DATA_BLOCK "LANGUAGE"   // DB4
TITLE = LANGUAGE
{ S7_Optimized_Access := 'FALSE' }
AUTHOR : oscat
FAMILY : CONSTANT
NAME : DBLANG
VERSION : 1.2
   VAR
      DEFAULT : Int := 1;   // 1=english, 2=german, 3=french
      LMAX : Int := 3;
      WEEKDAYS : Array[1..3, 1..7] of String[10];
      WEEKDAYS2 : Array[1..3, 1..7] of String[2];
      MONTHS : Array[1..3, 1..12] of String[10];
      MONTHS3 : Array[1..3, 1..12] of String[3];
      DIRS : Array[1..3, 0..15] of String[3];
   END_VAR
BEGIN
   WEEKDAYS[1,1] := 'Monday';
   WEEKDAYS[1,2] := 'Tuesday';
   WEEKDAYS[1,3] := 'Wednesday';
   WEEKDAYS[1,4] := 'Thursday';
   WEEKDAYS[1,5] := 'Friday';
   WEEKDAYS[1,6] := 'Saturday';
   WEEKDAYS[1,7] := 'Sunday';
   WEEKDAYS[2,1] := 'Montag';
   WEEKDAYS[2,2] := 'Dienstag';
   WEEKDAYS[2,3] := 'Mittwoch';
   WEEKDAYS[2,4] := 'Donnerstag';
   WEEKDAYS[2,5] := 'Freitag';
   WEEKDAYS[2,6] := 'Samstag';
   WEEKDAYS[2,7] := 'Sonntag';
   WEEKDAYS[3,1] := 'Lundi';
   WEEKDAYS[3,2] := 'Mardi';
   WEEKDAYS[3,3] := 'Mercredi';
   WEEKDAYS[3,4] := 'Jeudi';
   WEEKDAYS[3,5] := 'Vendredi';
   WEEKDAYS[3,6] := 'Samedi';
   WEEKDAYS[3,7] := 'Dimanche';
   WEEKDAYS2[1,1] := 'Mo';
   WEEKDAYS2[1,2] := 'Tu';
   WEEKDAYS2[1,3] := 'We';
   WEEKDAYS2[1,4] := 'Th';
   WEEKDAYS2[1,5] := 'Fr';
   WEEKDAYS2[1,6] := 'Sa';
   WEEKDAYS2[1,7] := 'Su';
   WEEKDAYS2[2,1] := 'Mo';
   WEEKDAYS2[2,2] := 'Di';
   WEEKDAYS2[2,3] := 'Mi';
   WEEKDAYS2[2,4] := 'Do';
   WEEKDAYS2[2,5] := 'Fr';
   WEEKDAYS2[2,6] := 'Sa';
   WEEKDAYS2[2,7] := 'So';
   WEEKDAYS2[3,1] := 'Lu';
   WEEKDAYS2[3,2] := 'Ma';
   WEEKDAYS2[3,3] := 'Me';
   WEEKDAYS2[3,4] := 'Je';
   WEEKDAYS2[3,5] := 'Ve';
   WEEKDAYS2[3,6] := 'Sa';
   WEEKDAYS2[3,7] := 'Di';
   MONTHS[1,1] := 'January';
   MONTHS[1,2] := 'February';
   MONTHS[1,3] := 'March';
   MONTHS[1,4] := 'April';
   MONTHS[1,5] := 'May';
   MONTHS[1,6] := 'June';
   MONTHS[1,7] := 'July';
   MONTHS[1,8] := 'August';
   MONTHS[1,9] := 'September';
   MONTHS[1,10] := 'October';
   MONTHS[1,11] := 'November';
   MONTHS[1,12] := 'December';
   MONTHS[2,1] := 'Januar';
   MONTHS[2,2] := 'Februar';
   MONTHS[2,3] := 'März';
   MONTHS[2,4] := 'April';
   MONTHS[2,5] := 'Mai';
   MONTHS[2,6] := 'Juni';
   MONTHS[2,7] := 'Juli';
   MONTHS[2,8] := 'August';
   MONTHS[2,9] := 'September';
   MONTHS[2,10] := 'Oktober';
   MONTHS[2,11] := 'November';
   MONTHS[2,12] := 'Dezember';
   MONTHS[3,1] := 'Janvier';
   MONTHS[3,2] := 'Février';
   MONTHS[3,3] := 'mars';
   MONTHS[3,4] := 'Avril';
   MONTHS[3,5] := 'Mai';
   MONTHS[3,6] := 'Juin';
   MONTHS[3,7] := 'Juillet';
   MONTHS[3,8] := 'Août';
   MONTHS[3,9] := 'Septembre';
   MONTHS[3,10] := 'Octobre';
   MONTHS[3,11] := 'Novembre';
   MONTHS[3,12] := 'Decembre';
   MONTHS3[1,1] := 'Jan';
   MONTHS3[1,2] := 'Feb';
   MONTHS3[1,3] := 'Mar';
   MONTHS3[1,4] := 'Apr';
   MONTHS3[1,5] := 'May';
   MONTHS3[1,6] := 'Jun';
   MONTHS3[1,7] := 'Jul';
   MONTHS3[1,8] := 'Aug';
   MONTHS3[1,9] := 'Sep';
   MONTHS3[1,10] := 'Oct';
   MONTHS3[1,11] := 'Nov';
   MONTHS3[1,12] := 'Dec';
   MONTHS3[2,1] := 'Jan';
   MONTHS3[2,2] := 'Feb';
   MONTHS3[2,3] := 'Mrz';
   MONTHS3[2,4] := 'Apr';
   MONTHS3[2,5] := 'Mai';
   MONTHS3[2,6] := 'Jun';
   MONTHS3[2,7] := 'Jul';
   MONTHS3[2,8] := 'Aug';
   MONTHS3[2,9] := 'Sep';
   MONTHS3[2,10] := 'Okt';
   MONTHS3[2,11] := 'Nov';
   MONTHS3[2,12] := 'Dez';
   MONTHS3[3,1] := 'Jan';
   MONTHS3[3,2] := 'Fev';
   MONTHS3[3,3] := 'Mar';
   MONTHS3[3,4] := 'Avr';
   MONTHS3[3,5] := 'Mai';
   MONTHS3[3,6] := 'Jun';
   MONTHS3[3,7] := 'Jul';
   MONTHS3[3,8] := 'Aou';
   MONTHS3[3,9] := 'Sep';
   MONTHS3[3,10] := 'Oct';
   MONTHS3[3,11] := 'Nov';
   MONTHS3[3,12] := 'Dec';
   DIRS[1,0] := 'N';
   DIRS[1,1] := 'NNE';
   DIRS[1,2] := 'NE';
   DIRS[1,3] := 'ENE';
   DIRS[1,4] := 'E';
   DIRS[1,5] := 'ESE';
   DIRS[1,6] := 'SE';
   DIRS[1,7] := 'SSE';
   DIRS[1,8] := 'S';
   DIRS[1,9] := 'SSW';
   DIRS[1,10] := 'SW';
   DIRS[1,11] := 'WSW';
   DIRS[1,12] := 'W';
   DIRS[1,13] := 'WNW';
   DIRS[1,14] := 'NW';
   DIRS[1,15] := 'NNW';
   DIRS[2,0] := 'N';
   DIRS[2,1] := 'NNO';
   DIRS[2,2] := 'NO';
   DIRS[2,3] := 'ONO';
   DIRS[2,4] := 'O';
   DIRS[2,5] := 'OSO';
   DIRS[2,6] := 'SO';
   DIRS[2,7] := 'SSO';
   DIRS[2,8] := 'S';
   DIRS[2,9] := 'SSW';
   DIRS[2,10] := 'SW';
   DIRS[2,11] := 'WSW';
   DIRS[2,12] := 'W';
   DIRS[2,13] := 'WNW';
   DIRS[2,14] := 'NW';
   DIRS[2,15] := 'NNW';
   DIRS[3,0] := 'N';
   DIRS[3,1] := 'NNO';
   DIRS[3,2] := 'NO';
   DIRS[3,3] := 'ONO';
   DIRS[3,4] := 'O';
   DIRS[3,5] := 'OSO';
   DIRS[3,6] := 'SO';
   DIRS[3,7] := 'SSO';
   DIRS[3,8] := 'S';
   DIRS[3,9] := 'SSW';
   DIRS[3,10] := 'SW';
   DIRS[3,11] := 'WSW';
   DIRS[3,12] := 'W';
   DIRS[3,13] := 'WNW';
   DIRS[3,14] := 'NW';
   DIRS[3,15] := 'NNW';
END_DATA_BLOCK

DATA_BLOCK "CONSTANTS"   // DB6
TITLE = CONSTANTS
{ S7_Optimized_Access := 'FALSE' }
AUTHOR : oscat
FAMILY : CONSTANT
NAME : CONSTANT
VERSION : 1.0
   VAR
      STRING_LENGTH : Int := 250;
      LIST_LENGTH : Int := 250;
   END_VAR
BEGIN
END_DATA_BLOCK

DATA_BLOCK "TEMP"   // DB7
TITLE = temporary Strings
{ S7_Optimized_Access := 'FALSE' }
AUTHOR : dalbi
FAMILY : xS7
NAME : DBTEMP
VERSION : 1.1
   VAR
      STR1 : String[254];
      STR2 : String[254];
      STR3 : String[254];
      TEMP : String[254];
   END_VAR
BEGIN
END_DATA_BLOCK

FUNCTION_BLOCK "MESSAGE_4R"   // FB34, SCL
TITLE = MESSAGE_4R
{ S7_Optimized_Access := 'FALSE' }
AUTHOR : hugo
FAMILY : STRINGS
NAME : MESSG4R
VERSION : 1.1
// this function generates a rotation meassage with up to 4 strings.
// on each rising edge of EN the next message in line will be displayed.
// when EN stays high longer then one cycle, the next message will be displayed automatically after the time T1 is elapsed.
// the output MX is the generated message and CX is a counter 0..3 signaling the current message displayed.
// the displayed messages are 0 .. MM.
// 
// uses: INC1 [FC53]
   VAR_INPUT
      M0 : String[254];
      M1 : String[254];
      M2 : String[254];
      M3 : String[254];
      MM : Int := 3;
      ENQ : Bool := TRUE;
      CLK : Bool := TRUE;
      T1 : Time := T#3S;
   END_VAR
   VAR_OUTPUT
      MX : String[254];
      MN : Int;
      TR : Bool;
   END_VAR
   VAR
      _timer : TON;
      edge : Bool;
   END_VAR
BEGIN


   (* check for rising edge on EN *)
   #TR := FALSE;
   IF #ENQ THEN
       IF (NOT #edge AND #CLK) OR #_timer.Q THEN
               #MN := "INC1"(N:=#MM,X:=#MN);
               #TR := TRUE;
               #_timer.IN := FALSE;
               CASE #MN OF
                   0 : #MX BLKMOV #M0;
                   1 : #MX BLKMOV #M1;
                   2 : #MX BLKMOV #M2;
                   3 : #MX BLKMOV #M3;
               END_CASE;
       END_IF;
       #edge := #CLK;
       #_timer( IN := #CLK, PT := #T1);
   ELSE
       #MX := '';
       #MN := 0;
   END_IF;




   (* revision history
   hm  8. oct. 2008    rev 1.0
       original version

   hm  27. oct. 2008   rev 1.1
       changed _INC to INC1

   *)
END_FUNCTION_BLOCK

FUNCTION_BLOCK "MESSAGE_8"   // FB35, SCL
TITLE = MESSAGE_8
{ S7_Optimized_Access := 'FALSE' }
AUTHOR : hugo
FAMILY : STRINGS
NAME : MESSAGE8
VERSION : 1.1
// this function generates one out of 4 messages specified by S1 .. S8.
// the selected message will be presented at the output M.
// In1 has higher priority then In2 which has higher priority then IN3 and in8 has the lowest priority.
   VAR_INPUT
      IN1 : Bool;
      IN2 : Bool;
      IN3 : Bool;
      IN4 : Bool;
      IN5 : Bool;
      IN6 : Bool;
      IN7 : Bool;
      IN8 : Bool;
      S1 : String[254];
      S2 : String[254];
      S3 : String[254];
      S4 : String[254];
      S5 : String[254];
      S6 : String[254];
      S7 : String[254];
      S8 : String[254];
   END_VAR
   VAR_OUTPUT
      "M" : String[254];
   END_VAR
BEGIN


     (* check if an alarm is present if yes set the output M otherwise clear M *)
     IF #IN1 THEN
       #"M" BLKMOV #S1;
     ELSIF #IN2 THEN
       #"M" BLKMOV #S2;
     ELSIF #IN3 THEN
       #"M" BLKMOV #S3;
     ELSIF #IN4 THEN
       #"M" BLKMOV #S4;
     ELSIF #IN5 THEN
       #"M" BLKMOV #S5;
     ELSIF #IN6 THEN
       #"M" BLKMOV #S6;
     ELSIF #IN7 THEN
       #"M" BLKMOV #S7;
     ELSIF #IN8 THEN
       #"M" BLKMOV #S8;
     ELSE
       #"M" := '';
     END_IF;

   (* revision history
   hm  26.12.2007      rev 1.0
       original version

   hm  29. mar. 2008   rev 1.1
       changed STRING to STRING(STRING_LENGTH)
   *)
END_FUNCTION_BLOCK

FUNCTION_BLOCK "TICKER"   // FB36, SCL
TITLE = TICKER
{ S7_Optimized_Access := 'FALSE' }
AUTHOR : hugo
FAMILY : STRINGS
NAME : TICKER
VERSION : 1.2
// Ticker sends a substring of text with length N every TD Milliseconds to generate a ticker. 
//  
// uses: MID [FC26]
   VAR_INPUT
      N : Int;
      PT : Time;
   END_VAR
   VAR_OUTPUT
      Display : String[254];
   END_VAR
   VAR_IN_OUT
      Text : String[254];
   END_VAR
   VAR
      delay : TP;
      "step" : Int;
   END_VAR
   VAR_TEMP
      tText : String[254];
      _Text AT tText : Struct
         length : Byte;
         act_length : Byte;
         str : Array[1..254] of Byte;
      END_STRUCT;
   END_VAR
BEGIN


   #tText := #Text; 

   (* generate next ticker when delay is low *)
   IF #N < BYTE_TO_INT(#_Text.act_length) THEN
       IF NOT #delay.Q THEN
         (* increase step for next tick *)
         #"step" := #"step" + 1;
         IF #"step" > BYTE_TO_INT(#_Text.act_length) THEN #"step" := 1; END_IF;
         (* extract dispay from text *)
         #Display := MID(IN:=#tText,L:=#N,P:=#"step");
         (* set delay timer for next tick *)
         #delay(IN := TRUE, PT := #PT);
       ELSE;
         (* execute delay timer *)
         #delay.IN := FALSE;
       END_IF;
   ELSE
       #Display BLKMOV #tText;
   END_IF;


   (* revision history
   hm  4. dec. 2007    rev 1.0
       original version

   hm  15. dec. 2007   rev 1.1
       step now starts at 1 instaed of 0

   hm  29. mar. 2008   rev 1.2
       changed STRING to STRING(STRING_LENGTH)
   *)
END_FUNCTION_BLOCK

FUNCTION "INC1" : Int   // FC53, SCL
TITLE = INC1
{ S7_Optimized_Access := 'FALSE' }
AUTHOR : hugo
FAMILY : MATH
NAME : INC1
VERSION : 1.2
// This is a increment function which increments the variable X by 1 and if M is reached, it begins with 0 again.
// _inc1(3,X) will generate 0,1,2,3,0,1,.....
   VAR_INPUT
      X : Int;
      N : Int;
   END_VAR
BEGIN


   IF #X >= #N - 1 THEN
       #INC1 := 0;
   ELSE
       #INC1 := #X + 1;
   END_IF;


   (* this elegant version is 50% slower
   INC1 := X := (x + 1) MOD N;
   *)



   (* revision history
   hm  13. oct. 2008   rev 1.0
       original version

   hm  22. oct. 2008   rev 1.1
       added statement to return value for compatibility reasons

   hm  23. feb. 2009   rev 1.2
       when inc1 is called with X >= N inc will continue with 0
   *)
END_FUNCTION

FUNCTION "EXP10" : Real   // FC77, SCL
TITLE = EXP10
{ S7_Optimized_Access := 'FALSE' }
AUTHOR : hugo
FAMILY : MATH
NAME : exp10
VERSION : 1.0
// this function calculates the exponent to the basis 10
// exp10(3) = 1000
   VAR_INPUT
      X : Real;
   END_VAR
BEGIN


     #EXP10 := EXP(#X * 2.30258509299405);

   (* revision history
   hm  2. dec 2007    rev 1.0
     original version

   *)
END_FUNCTION

FUNCTION "EXPN" : Real   // FC78, SCL
TITLE = EXPN
{ S7_Optimized_Access := 'FALSE' }
AUTHOR : hugo
FAMILY : MATH
NAME : EXPN
VERSION : 1.2
// this function calculates X to the power of N (Y = X^N) whilke N is an integer
// especially on CPU's without a floating point unit this algorythm is about 30 times faster then the IEC standard EXPT() Function
   VAR_INPUT
      X : Real;
      N : Int;
   END_VAR
   VAR_TEMP
      tempN : Int;
      _tempN AT tempN : Array[0..15] of Bool;
      tempX : Real;
      sign : Bool;
   END_VAR
BEGIN


   #tempN := #N;
   #tempX := #X;

   #sign := #_tempN[7]; //N.15
   #tempN := ABS(#tempN);
   IF #_tempN[8] THEN #EXPN := #tempX; ELSE #EXPN := 1.0; END_IF;
   #tempN := WORD_TO_INT(SHR(IN:=INT_TO_WORD(#tempN),N:=1));
   WHILE #tempN > 0 DO
      #tempX := #tempX * #tempX;
      IF #_tempN[8] THEN #EXPN := #EXPN * #tempX; END_IF;
      #tempN := WORD_TO_INT(SHR(IN:=INT_TO_WORD(#tempN),N:=1));
   END_WHILE;
   IF #sign THEN #EXPN := 1.0 / #EXPN; END_IF;


   (* revision history
   hm  4. dec 2007 rev 1.0
       original version

   hm  22. oct. 2008   rev 1.1
       optimized code

   hm  10. mar. 2009   rev 1.2
       removed nested comments
       real constants updated to new systax using dot

   *)
END_FUNCTION

FUNCTION "DAY_OF_MONTH" : Int   // FC178, SCL
TITLE = DAY_OF_MONTH
{ S7_Optimized_Access := 'FALSE' }
AUTHOR : hugo
FAMILY : TIDT
NAME : DAYOMON
VERSION : 2.1
// returns the day OF month from any DATE
// 
// uses: DAY_OF_YEAR [FC180]
//       YEAR_BEGIN [FC217] 
//       YEAR_OF_DATE [FC219] 
//       LEAP_OF_DATE [FC193]
//       LEAP_YEAR [FC194]
   VAR_INPUT
      IDATE : Date;
   END_VAR
   VAR_TEMP
      leap : Int;
   END_VAR
BEGIN


   (* calculate the day in the year *)
   #DAY_OF_MONTH := "DAY_OF_YEAR"(#IDATE);
   (* leap will be set to one for a leap year *)
   #leap := BOOL_TO_INT("LEAP_OF_DATE"(#IDATE));
   (* if leap year deduct one from the days of the year *)
   #DAY_OF_MONTH := #DAY_OF_MONTH - #leap;
   (* search if we are in month december to march ? *)
   IF #DAY_OF_MONTH > "MTH_OFS9" THEN
       IF #DAY_OF_MONTH > "MTH_OFS11" THEN
           IF #DAY_OF_MONTH > "MTH_OFS12" THEN
               #DAY_OF_MONTH := #DAY_OF_MONTH - "MTH_OFS12";
           ELSE
               #DAY_OF_MONTH := #DAY_OF_MONTH - "MTH_OFS11";
           END_IF;
       ELSE
           IF #DAY_OF_MONTH > "MTH_OFS10" THEN
               #DAY_OF_MONTH := #DAY_OF_MONTH - "MTH_OFS10";
           ELSE
               #DAY_OF_MONTH := #DAY_OF_MONTH - "MTH_OFS9";
           END_IF;
       END_IF;
   ELSIF #DAY_OF_MONTH > "MTH_OFS5" THEN
       IF #DAY_OF_MONTH > "MTH_OFS7" THEN
           IF #DAY_OF_MONTH > "MTH_OFS8" THEN
               #DAY_OF_MONTH := #DAY_OF_MONTH - "MTH_OFS8";
           ELSE
               #DAY_OF_MONTH := #DAY_OF_MONTH - "MTH_OFS7";
           END_IF;
       ELSE
           IF #DAY_OF_MONTH > "MTH_OFS6" THEN
               #DAY_OF_MONTH := #DAY_OF_MONTH - "MTH_OFS6";
           ELSE
               #DAY_OF_MONTH := #DAY_OF_MONTH - "MTH_OFS5";
           END_IF;
       END_IF;
   ELSIF #DAY_OF_MONTH > "MTH_OFS3" THEN
       IF #DAY_OF_MONTH > "MTH_OFS4" THEN
           #DAY_OF_MONTH := #DAY_OF_MONTH - "MTH_OFS4";
       ELSE
           #DAY_OF_MONTH := #DAY_OF_MONTH - "MTH_OFS3";
       END_IF;
   ELSE
       (* since now we must be in february or january we need to add leap again *)
       #DAY_OF_MONTH := #DAY_OF_MONTH + #leap;
       IF #DAY_OF_MONTH > "MTH_OFS2" THEN #DAY_OF_MONTH := #DAY_OF_MONTH - "MTH_OFS2"; END_IF;
       (* since nothing was true before, day_of_month must already be good *)
   END_IF;


   (*
   Revision history

   hm 22.1.2007        rev 1.1
       deleted unused variable day_in_year and day_in_year_begin

   hm  1. okt 2007 rev 1.2
       changed code to use day_of_year and leap_of_date
       added compatibility to STEP7

   hm  8. oct 2007 rev 1.3
       deleted unused variable yr

   hm  8. jan 2008 rev 1.4
       improved performance

   hm  25. oct. 2008   rev 2.0
       new code using setup constants

   hm  10. mar. 2009   rev 2.1
       removed nested comments

   *)
END_FUNCTION

FUNCTION "DAY_OF_WEEK" : Int   // FC179, SCL
TITLE = DAY_OF_WEEK
{ S7_Optimized_Access := 'FALSE' }
AUTHOR : hugo
FAMILY : TIDT
NAME : DWEEK
VERSION : 1.4
// calculates the weekday of a week according to ISO8601   
// monday = 1 ..... sunday = 7
   VAR_INPUT
      IDATE : Date;
   END_VAR
BEGIN


     #DAY_OF_WEEK := DINT_TO_INT((T_CONV(#IDATE)+7308) MOD 7)+1;

   (* 
   weekday := DWORD_TO_INT((DATE_TO_DWORD(idate)/86400+3) MOD 7) + 1;
   *)


   (* revision history
   hm  21.8.06         rev 1.1
       corrected a miscalculation

   hm  23.12.2007      rev 1.2
       correction for step7

   hm  7. apr. 2008    rev 1.3
       deleted unused step7 code

   hm  7. oct. 2008    rev 1.4
       changed name of function from weekday to day_of_week

   *)
END_FUNCTION

FUNCTION "DAY_OF_YEAR" : Int   // FC180, SCL
TITLE = DAY_OF_YEAR
{ S7_Optimized_Access := 'FALSE' }
AUTHOR : hugo
FAMILY : TIDT
NAME : DAYOYEAR
VERSION : 1.4
// calculates the day of the year
// 
// uses: DATE_DINT [FC405]
   VAR_INPUT
      idate : Date;
   END_VAR
BEGIN


   #DAY_OF_YEAR := DINT_TO_INT(("DATE_DINT"(#idate) / 86400) MOD 1461);
   IF #DAY_OF_YEAR > 729 THEN
     IF #DAY_OF_YEAR > 1095 THEN #DAY_OF_YEAR := #DAY_OF_YEAR - 1095; ELSE #DAY_OF_YEAR := #DAY_OF_YEAR - 729; END_IF;
   ELSIF #DAY_OF_YEAR > 364 THEN
     #DAY_OF_YEAR := #DAY_OF_YEAR - 364;
   ELSE
     #DAY_OF_YEAR := #DAY_OF_YEAR + 1;
   END_IF;

   //  day_of_year := DINT_TO_INT((DATE_TO_DINT(idate) - DATE_TO_DINT(year_begin(year_of_date(idate))))) + 1;

   (*
   DAY_OF_YEAR := DWORD_TO_INT((DATE_TO_DWORD(idate) - DATE_TO_DWORD(YEAR_BEGIN(YEAR_OF_DATE(idate)))) / 86400) + 1;
   *)


   (* revivision history
   hm  4. aug. 2007    rev 1.0
     original version

   hm  1. oct. 2007    rev 1.1
     added compatibility to STEP7

   hm  4. jan. 2008    rev 1.2
     changed code for better performance

   hm  7. oct. 2008    rev 1.3
     changed name of function year to year_of_date

   hm  28. jan. 2011 rev 1.4
     improved code
   *)
END_FUNCTION

FUNCTION "HOUR" : Int   // FC187, SCL
TITLE = HOUR
{ S7_Optimized_Access := 'FALSE' }
AUTHOR : hugo
FAMILY : TIDT
NAME : HOUR
VERSION : 1.1
// extracts the hour of a Time_of_day
   VAR_INPUT
      itod : Time_Of_Day;
   END_VAR
BEGIN


     #HOUR := DINT_TO_INT(T_CONV(#itod)/3600000);

   (* change history
   hm 4. aug 2006  rev 1.0
     original version

   hm 2.10.2006   rev 1.1
     changed name of input to itod

   *)
END_FUNCTION

FUNCTION "LEAP_OF_DATE" : Bool   // FC193, SCL
TITLE = LEAP_OF_DATE
{ S7_Optimized_Access := 'FALSE' }
AUTHOR : hugo
FAMILY : TIDT
NAME : LEAPODAT
VERSION : 1.3
// leap_year is true if the tested year is a leap year  
// 
// uses: DATE_DINT [FC405]
   VAR_INPUT
      idate : Date;
   END_VAR
BEGIN


   #LEAP_OF_DATE := SHL(IN:=DINT_TO_DWORD((("DATE_DINT"(#idate) + 43200) / 31557600)),N:=30) = 16#80000000;


   (* change history

   2.10.2006   rev 1.1
   the function now calls leap_year to accomodate further accuracy.
   the function now works for any year from 1970 to 2100

   8. jan 2008   rev 1.2
     improved code for better performance

   28. jan. 2011 rev 1.3
     improved performance
   *)
END_FUNCTION

FUNCTION "MINUTE" : Int   // FC197, SCL
TITLE = MINUTE
{ S7_Optimized_Access := 'FALSE' }
AUTHOR : hugo
FAMILY : TIDT
NAME : MINUTE
VERSION : 1.1
// extracts the minutes out of TOD truncating the ceconds
   VAR_INPUT
      itod : Time_Of_Day;
   END_VAR
BEGIN


     #MINUTE := DINT_TO_INT(T_CONV(#itod)/60000 - T_CONV(#itod)/3600000 * 60);


   (* change history

   2.10.2006 changes name of input to itod

   *)
END_FUNCTION

FUNCTION "MONTH_OF_DATE" : Int   // FC202, SCL
TITLE = MONTH_OF_DATE
{ S7_Optimized_Access := 'FALSE' }
AUTHOR : hugo
FAMILY : TIDT
NAME : MONTH
VERSION : 1.3
// returns the month of a date  
// 
// uses: DAY_OF_YEAR [FC180]
//       YEAR_BEGIN [FC217] 
//       YEAR_OF_DATE [FC219] 
//       LEAP_OF_DATE [FC193]
//       LEAP_YEAR [FC194]
   VAR_INPUT
      IDATE : Date;
   END_VAR
BEGIN


   #MONTH_OF_DATE := "DAY_OF_YEAR"(#IDATE);
   IF #MONTH_OF_DATE < 32 THEN
       #MONTH_OF_DATE := 1;
   ELSIF "LEAP_OF_DATE"(#IDATE) THEN
       #MONTH_OF_DATE := (#MONTH_OF_DATE * 53 + 1668) / 1623;
   ELSE
       #MONTH_OF_DATE := (#MONTH_OF_DATE * 53 + 1700) / 1620;
   END_IF;


   (* code for rev 1.2
   MONTH_OF_DATE := DAY_OF_YEAR(IDATE);
   IF LEAP_OF_DATE(IDATE) THEN
       CASE MONTH_OF_DATE OF
           1..31   :   MONTH_OF_DATE := 1;
           32..60  :   MONTH_OF_DATE := 2;
           61..91  :   MONTH_OF_DATE := 3;
           92..121 :   MONTH_OF_DATE := 4;
           122..152:   MONTH_OF_DATE := 5;
           153..182:   MONTH_OF_DATE := 6;
           183..213:   MONTH_OF_DATE := 7;
           214..244:   MONTH_OF_DATE := 8;
           245..274:   MONTH_OF_DATE := 9;
           275..305:   MONTH_OF_DATE := 10;
           306..335:   MONTH_OF_DATE := 11;
           336..366:   MONTH_OF_DATE := 12;
       END_CASE;
   ELSE
       CASE MONTH_OF_DATE OF
           1..31   :   MONTH_OF_DATE := 1;
           32..59  :   MONTH_OF_DATE := 2;
           60..90  :   MONTH_OF_DATE := 3;
           91..120 :   MONTH_OF_DATE := 4;
           121..151:   MONTH_OF_DATE := 5;
           152..181:   MONTH_OF_DATE := 6;
           182..212:   MONTH_OF_DATE := 7;
           213..243:   MONTH_OF_DATE := 8;
           244..273:   MONTH_OF_DATE := 9;
           274..304:   MONTH_OF_DATE := 10;
           305..334:   MONTH_OF_DATE := 11;
           335..365:   MONTH_OF_DATE := 12;
       END_CASE;
   END_IF;
   *)


   (* revision history
   hm  1. aug 2006 rev 1.0
       original version    

   hm  1. okt 2007 rev 1.1
       replaced old code (string conversion) with mathematics
       the execution time is now multiple times faster.

   hm  7. oct. 2008    rev 1.2
       changed name of function from month to MONTH_OF_DATE

   hm  27. mar. 2009   rev 1.3
       new improved code

   *)
END_FUNCTION

FUNCTION "SECOND" : Real   // FC210, SCL
TITLE = SECOND
{ S7_Optimized_Access := 'FALSE' }
AUTHOR : hugo
FAMILY : TIDT
NAME : SEC
VERSION : 1.1
// returns the seconds and milliseconds as real of TOD
   VAR_INPUT
      itod : Time_Of_Day;
   END_VAR
BEGIN


     #SECOND := DINT_TO_REAL(T_CONV(#itod) - T_CONV(#itod)/60000 * 60000)/1000;



   (* change history

   2.10.2006 changes name of input to itod

   *)
END_FUNCTION

FUNCTION "SET_DT" : Date_And_Time   // FC214, SCL
TITLE = SET_DT
{ S7_Optimized_Access := 'FALSE' }
AUTHOR : hugo
FAMILY : TIDT
NAME : SET_DT
VERSION : 1.5
// creates a date output from year, month and day of month
// year must be in the form of 4 digits ie 2006 or 1977.
   VAR_INPUT
      year : Int;
      month : Int;
      day : Int;
      hour : Int;
      minute : Int;
      second : Int;
   END_VAR
   VAR_TEMP
      tDT : Date_And_Time;
      _DT AT tDT : Array[0..7] of Byte;
      t_year : Int;
   END_VAR
BEGIN


     //set_DT := DWORD_TO_DT(DATE_TO_DWORD(set_Date(year, month, day)) + second + minute * 60 + INT_TO_DWORD(hour) * 3600);

     #t_year := #year - 1900;

     IF #t_year > 99 THEN 
       #t_year := #year - 2000; 
     END_IF;

     #_DT[0] := WORD_TO_BYTE(INT_TO_BCD16(#t_year));   // year
     #_DT[1] := WORD_TO_BYTE(INT_TO_BCD16(#month));    // month
     #_DT[2] := WORD_TO_BYTE(INT_TO_BCD16(#day));      // day
     #_DT[3] := WORD_TO_BYTE(INT_TO_BCD16(#hour));     // hour
     #_DT[4] := WORD_TO_BYTE(INT_TO_BCD16(#minute));   // minute
     #_DT[5] := WORD_TO_BYTE(INT_TO_BCD16(#second));   // second

     #SET_DT := #tDT;

   (* revision history
   hm  4. aug. 2006        rev 1.0
       original version

   hm      19 sep. 2007    rev 1.1
       use function leap_year to calculate leap year, more exceptions are handled

   hm      1. okt 2007     rev 1.2
       added step7 compatibility
       call function set_date

   hm      8. oct 2007     rev 1.3
       deleted unused variables count and leap

   hm      1. 11 2007      rev 1.4
       converted hour type integer to dword in calculation to avoid overrun on möller ecp4

   hm      16. mar 2008    rev 1.5
       added type conversions to avoid warnings under codesys 3.0
   *)
END_FUNCTION

FUNCTION "YEAR_OF_DATE" : Int   // FC219, SCL
TITLE = YEAR_OF_DATE
{ S7_Optimized_Access := 'FALSE' }
AUTHOR : hugo
FAMILY : TIDT
NAME : YEAR
VERSION : 1.4
// returs the year of a date  
// the function works for dates from 1990 - 2100
   VAR_INPUT
      IDATE : Date;
   END_VAR
BEGIN


   #YEAR_OF_DATE := DINT_TO_INT(((100 * T_CONV(#IDATE)) + 50) / 36525) + 1990;  

   (*
   year := DWORD_TO_INT((DATE_TO_DWORD(idate)+43200) / 31557600 + 1970);
   *)

   (* code used prior to rev 1.1
   year := DWORD_TO_INT((DATE_TO_DWORD(idate)/864+71954300)/36525);
   *)

   (* revision history
   hm  4. aug 2006     rev 1.0
       original version

   hm  1. okt 2007     rev 1.1
       corrected error in algorithm
       adjustment for S7 compatibility

   hm  23.12.2007      rev 1.2
       changed code for better performance

   hm  7. apr. 2008    rev 1.3
       deleted unused step7 code

   hm  7. oct. 2008    rev 1.4
       reneamed function (year) to year_of_date

   *)
END_FUNCTION

FUNCTION "BIN_TO_BYTE" : Byte   // FC220, SCL
TITLE = BIN_TO_BYTE
{ S7_Optimized_Access := 'FALSE' }
AUTHOR : hugo
FAMILY : STRINGS
NAME : BIN2BY
VERSION : 1.2
// BINARY_TO_byte converts a binary string into a byte.
   VAR_INPUT
      BIN : String[254];
      _BIN AT BIN : Struct
         length : Byte;
         act_length : Byte;
         str : Array[1..12] of Byte;
      END_STRUCT;
   END_VAR
   VAR_TEMP
      pt : Int;   // pt : POINTER TO BYTE;
      i : Int;
      X : Byte;
      stop : Int;
   END_VAR
BEGIN


   #pt := 1;    //ADR(bin);
   #stop := BYTE_TO_INT(#_BIN.act_length);    //LEN(bin);
   FOR #i := 1 TO #stop DO
     (* read the first character and subtract 48 to get value in decimal 0 = 48 *)
     #X := #_BIN.str[#pt];
     (* calculate the value of the digit *)
     IF #X = 48 THEN
       #BIN_TO_BYTE := SHL(IN:=#BIN_TO_BYTE, N:=1);
     ELSIF #X = 49 THEN
       #BIN_TO_BYTE := SHL(IN:=#BIN_TO_BYTE, N:=1) OR 1;
     END_IF;
     #pt := #pt + 1;
   END_FOR;


   (* revision histroy
   hm  18. jun. 2008 rev 1.0
     original release

   hm  20. sep. 2008 rev 1.1
     changed length of input string from 20 to 12

   hm  26. jul. 2009 rev 1.2
     optimized code
   *)
END_FUNCTION

FUNCTION "BIN_TO_DWORD" : DWord   // FC221, SCL
TITLE = BIN_TO_DWORD
{ S7_Optimized_Access := 'FALSE' }
AUTHOR : hugo
FAMILY : STRINGS
NAME : BIN2DW
VERSION : 1.2
// BINARY_TO_DWORD converts a binary string into a dword.
   VAR_INPUT
      BIN : String[254];
      _BIN AT BIN : Struct
         length : Byte;
         act_length : Byte;
         str : Array[1..40] of Byte;
      END_STRUCT;
   END_VAR
   VAR_TEMP
      pt : Int;   // pt : POINTER TO BYTE;
      i : Int;
      X : Byte;
      stop : Int;
   END_VAR
BEGIN


   #pt := 1;    //ADR(bin);
   #stop := BYTE_TO_INT(#_BIN.act_length);     //LEN(bin);
   FOR #i := 1 TO #stop DO
     (* read the first character and subtract 48 to get value in decimal 0 = 48 *)
     #X := #_BIN.str[#pt];
     (* calculate the value of the digit *)
     IF BYTE_TO_INT(#X) = 48 THEN
       #BIN_TO_DWORD := SHL(IN:=#BIN_TO_DWORD, N:=1);
     ELSIF BYTE_TO_INT(#X) = 49 THEN
       #BIN_TO_DWORD := SHL(IN:=#BIN_TO_DWORD, N:=1) OR 1;
     END_IF;
     #pt := #pt + 1;
   END_FOR;


   (* revision histroy
   hm  18. jun. 2008 rev 1.0
     original release

   hm  20. sep. 2008 rev 1.1
     changed length of input dtring from 20 to 40

   hm  26. jul 2009  rev 1.2
     optimized code
   *)
END_FUNCTION

FUNCTION "BYTE_TO_STRB" : String[254]   // FC222, SCL
TITLE = BYTE_TO_STRB
{ S7_Optimized_Access := 'FALSE' }
AUTHOR : hugo
FAMILY : STRINGS
NAME : BYTSTRB
VERSION : 1.3
// BYTE_TO_STRINGB converts a Byte to a String of Bits represented by '0' and '1' s.
// The lowest order bit will be on the right and the high order bit on the left.
   VAR_INPUT
      IN : Byte;
   END_VAR
   VAR_TEMP
      i : Int;
      pt : Int;   // pt : POINTER TO BYTE;
      str : String[8];
      _str AT str : Struct
         length : Byte;
         act_length : Byte;
         str : Array[1..8] of Byte;
      END_STRUCT;
      tIN : Byte;
      _IN AT tIN : Array[0..7] of Bool;
   END_VAR
BEGIN


   #str := #BYTE_TO_STRB;
   #tIN := #IN;

   (* pointer für die ausgabe ermitteln *)
   #pt := 1;    //ADR(BYTE_TO_STRB);
   (* die 8 ausgabecharacter ermitteln und schreiben *)
   FOR #i := 1 TO 8 DO
       #_str.str[#pt] := INT_TO_BYTE(BYTE_TO_INT(BOOL_TO_BYTE(#_IN[7])) + 48); 
       #tIN := SHL(IN:=#tIN,N:=1);
       #pt := #pt + 1;
   END_FOR;

   (* der ausgabestring muss noch mit 8 abgeschlossen werden *)
   #_str.act_length := 8;
   #BYTE_TO_STRB := #str;

   (* code before rev 1.1
   FOR i := 1 TO 8 DO
       IF in.0 = 0 THEN temp := CONCAT('0', temp); ELSE temp := CONCAT('1', temp); END_IF;
       in := SHR(in, 1);
   END_FOR;
   BYTE_TO_STRB := temp;
   *)


   (* revision history

   hm      9.6.2007    rev 1.0     
       original version 

   hm  15. dec 2007    rev 1.1
       inprooved code for higher performance

   hm  29. mar. 2008   rev 1.2
       changed STRING to STRING(8)

   hm  20. jun. 2008   rev 1.3
       performance improvement

   *)
END_FUNCTION

FUNCTION "BYTE_TO_STRH" : String[254]   // FC223, SCL
TITLE = BYTE_TO_STRH
{ S7_Optimized_Access := 'FALSE' }
AUTHOR : hugo
FAMILY : STRINGS
NAME : BYTSTRH
VERSION : 1.3
// BYTE_TO_STRINGH converts a Byte to a String of Hexadecimal represented by '0' .. '9' and 'A' .. 'F'.
// The lowest order Character will be on the right and the high order Character on the left.
   VAR_INPUT
      IN : Byte;
   END_VAR
   VAR_TEMP
      temp : Byte;
      PT : Int;   // PT : POINTER TO BYTE;
      str : String[2];
      _str AT str : Struct
         length : Byte;
         act_length : Byte;
         str : Array[1..2] of Byte;
      END_STRUCT;
   END_VAR
BEGIN


   #str := #BYTE_TO_STRH;

   (* read pointer to output string *)
   #PT := 1;    //ADR(BYTE_TO_STRH);
   (* calculate high order hex value *)
   #temp := SHR(IN:=#IN,N:=4);
   (* convert value to hex character *)
   IF BYTE_TO_INT(#temp) <= 9 THEN #temp := INT_TO_BYTE(BYTE_TO_INT(#temp) + 48); ELSE #temp := INT_TO_BYTE(BYTE_TO_INT(#temp) + 55); END_IF;
   (* write friat character to output string *)
   #_str.str[#PT] := #temp;
   (* calculate low order hex value *)
   #temp := #IN AND 2#00001111;
   IF BYTE_TO_INT(#temp) <= 9 THEN #temp := INT_TO_BYTE(BYTE_TO_INT(#temp) + 48); ELSE #temp := INT_TO_BYTE(BYTE_TO_INT(#temp) + 55); END_IF;
   (* increment pointer and wirte low order character *)
   #PT := #PT + 1;
   #_str.str[#PT] := #temp;
   (* set pointer at the end of the output string and close the string with 2 *)
   #PT := #PT + 1;
   #_str.act_length := 2;
   #BYTE_TO_STRH := #str;

   (* code before rev 1.2
   FOR i := 1 TO 2 DO
       X := in AND 2#1111;
       IF X <= 9 THEN X := X + 48; ELSE X := X + 55; END_IF;
       Cx := CHR(X);
       temp := CONCAT(Cx, temp);
       in := SHR(in,4);
   END_FOR;
   BYTE_TO_STRH := temp;
   *)

   (* revision history

   hm  9.6.2007        rev 1.0     
       original version 

   hm  11.9.2007       rev 1.1     
       changed coding for compatibility with twincat, under twincat concat cannot have a function as argument.   

   hm  15 dec 2007     REV 1.2
       changed code for higher performance

   hm  29. mar. 2008   rev 1.3
       changed STRING to STRING(2)
   *)
END_FUNCTION

FUNCTION "CAPITALIZE" : String[254]   // FC224, SCL
TITLE = CAPITALIZE
{ S7_Optimized_Access := 'FALSE' }
AUTHOR : hugo
FAMILY : STRINGS
NAME : CAPITAL
VERSION : 1.1
// uppercase returns str while all letters a..z and ä,ö,ü are converted to uppercase
// 
// uses: SETUP [DB1]
//       TO_UPPER [FC284]
   VAR_INPUT
      str : String[254];
   END_VAR
   VAR_TEMP
      tCAPITALIZE : String[254];
      _CAPITALIZE AT tCAPITALIZE : Struct
         length : Byte;
         act_length : Byte;
         str : Array[1..254] of Byte;
      END_STRUCT;
      PT : Int;   // PT : POINTER TO BYTE;
      pos : Int;
      L : Int;
      first : Bool;
   END_VAR
BEGIN


   #first := TRUE;

   #PT := 1;    //ADR(CAPITALIZE);
   #tCAPITALIZE := #str;
   #L := BYTE_TO_INT(#_CAPITALIZE.act_length);   //LEN(str);
   FOR #pos := 1 TO #L DO
       IF #first THEN
           #_CAPITALIZE.str[#PT] := "TO_UPPER"(#_CAPITALIZE.str[#PT]);
       END_IF;
       (* remember in first if the next char needs to capitalized *)
       IF BYTE_TO_INT(#_CAPITALIZE.str[#PT]) = 32 THEN #first := TRUE; ELSE #first := FALSE; END_IF;
       #PT := #PT + 1;
   END_FOR;

   #CAPITALIZE := #tCAPITALIZE;

   (* revision histroy
   hm      4. mar 2008 rev 1.0
       original release

   hm  29. mar. 2008   rev 1.1
       changed STRING to STRING(STRING_LENGTH)
   *)
END_FUNCTION

FUNCTION "CHARCODE" : Byte   // FC225, SCL
TITLE = CHARCODE
{ S7_Optimized_Access := 'FALSE' }
AUTHOR : hugo
FAMILY : STRINGS
NAME : CHRCODE
VERSION : 1.2
// CHARCODE converts a HTML Character NAME INTO ITS code
// 'äuml' is convterted to ä
// 'euro' is converted to €
// 
// uses: SETUP [DB1]
//       CONCAT [FC2]
//       NE_STRNG [FC29]
//       LEN [FC21]
//       CODE [FC229]
//       FIND [FC11]
//       MID [FC26]
   VAR_INPUT
      STR : String[254];
   END_VAR
   VAR_TEMP
      tSTR : String[10];
      found : String[1];
      search : String[10];
      pos : Int;
      i : Int;
   END_VAR
BEGIN


   #tSTR := #STR;

   IF LEN(#tSTR) = 1 THEN
       #CHARCODE := "CODE"(STR:=#tSTR,POS:=1);
   ELSIF #tSTR <> '' THEN
       (* construct search string *)
       #search := CONCAT(IN1:='&',IN2:=#tSTR);
       #search := CONCAT(IN1:=#search, IN2:=';');
       WHILE #pos = 0 AND (#i < 4) DO
           #i := #i + 1;
           #pos := FIND(IN1:="SETUP".CHARNAMES[#i], IN2:=#search);
       END_WHILE;
       #found := MID(IN:="SETUP".CHARNAMES[#i], L:=1, P:=#pos - 1);
       #CHARCODE := "CODE"(STR:=#found, POS:=1);
   END_IF;

   (* revision history
   hm  13. may. 2008   rev 1.0
       original version

   hm  19. oct. 2008   rev 1.1
       changed setup constants

   hm  24. oct. 2008   rev 1.2
       optimized code
   *)
END_FUNCTION

FUNCTION "CHARNAME" : String[254]   // FC226, SCL
TITLE = CHARNAME
{ S7_Optimized_Access := 'FALSE' }
AUTHOR : hugo
FAMILY : STRINGS
NAME : CHRNAME
VERSION : 1.4
// CHARNAME converts a Character code into its HTML character name
// ä is convterted to 'äuml'
// € is converted to 'euro'
// 
// uses: SETUP [DB1]
//       CONCAT [FC2]
//       CHR_TO_STRING [FC227]
//       FIND [FC11]
//       MID [FC26]
//       LEFT [FC20]
   VAR_INPUT
      C : Byte;
   END_VAR
   VAR_TEMP
      search : String[254];
      pos : Int;
      tCHARNAME : String[10];
      i : Int;
   END_VAR
BEGIN


   #tCHARNAME := #CHARNAME;

   IF #C <> 0 THEN
       (* construct search string from code followed by $ sign, also clear charname string*)
       #tCHARNAME := "CHR_TO_STRING"(#C);
       #tCHARNAME := CONCAT(IN1:=#tCHARNAME,IN2:='&');
       #tCHARNAME := CONCAT(IN1:=';', IN2:=#tCHARNAME);
       WHILE #pos = 0 AND (#i < 4) DO
           #i := #i + 1;
           #pos := FIND(IN1:="SETUP".CHARNAMES[#i], IN2:=#tCHARNAME);
       END_WHILE;
       IF #pos > 0 THEN
           #tCHARNAME := MID(IN:="SETUP".CHARNAMES[#i], L:=10, P:=#pos + 3);
           (* search for end of name and truncate *)
           #pos := FIND(IN1:=#tCHARNAME, IN2:=';');
           #tCHARNAME := LEFT(IN:=#tCHARNAME,L:=#pos - 1);
       ELSE
           #tCHARNAME := "CHR_TO_STRING"(#C);
       END_IF;
   ELSE
       #tCHARNAME := '';
   END_IF;

   #CHARNAME := #tCHARNAME;


   (* revision history
   hm  13. may. 2008   rev 1.0
       original version

   hm  16. jun. 2008   rev 1.1
       changed nested call of concat for better compatibility

   hm  19. oct. 2008   rev 1.2
       changes setup constants

   hm  24. oct. 2008   rev 1.3
       new code for high performance

   hm  17. dec. 2008   rev 1.4
       changed function chr to chr_to_string
   *)
END_FUNCTION

FUNCTION "CHR_TO_STRING" : String[254]   // FC227, SCL
TITLE = CHR_TO_STRING
{ S7_Optimized_Access := 'FALSE' }
AUTHOR : hugo
FAMILY : STRINGS
NAME : CHRSTR
VERSION : 1.3
// CHR creates a character from a byte input and stuffs it in a one character length string.
   VAR_INPUT
      C : Byte;
   END_VAR
   VAR_TEMP
      tCHR : String[1];
      _CHR AT tCHR : Array[0..2] of Byte;
   END_VAR
BEGIN


   #_CHR[0] := 1;   (* length *)
   #_CHR[1] := 1;   (* actual length *)
   #_CHR[2] := #C; 
   #CHR_TO_STRING := #tCHR;

   (* revision history
   hm  16 jan 2007     rev 1.0
       original version

   hm  4. feb. 2008    rev 1.1
       return string would not be terminated properly

   hm  29. mar. 2008   rev 1.2
       changed STRING to STRING(1)

   hm  17. dec. 2008   rev 1.3
       changed name of function from chr to chr_to_string
   *)
END_FUNCTION

FUNCTION "CLEAN" : String[254]   // FC228, SCL
TITLE = CLEAN
{ S7_Optimized_Access := 'FALSE' }
AUTHOR : hugo
FAMILY : STRINGS
NAME : CLEAN
VERSION : 1.0
// Clean deletes all characters from a string except the ones specified in CX.
// 
// uses: LEN [FC21]
//       FIND [FC11]
//       MID [FC26]
//       DELETE [FC4]
   VAR_INPUT
      IN : String[254];
      CX : String[254];
   END_VAR
   VAR_TEMP
      tCLEAN : String[254];
      tCX : String[80];
      pos : Int;
      stop : Int;
   END_VAR
BEGIN


   #pos := 1;
   #tCLEAN := #IN;
   #tCX := #CX;

   (* copy input string *)
   //CLEAN := IN;
   #stop := LEN(#tCLEAN);
   WHILE #pos <= #stop DO
       IF FIND(IN1:=#tCX,IN2:=MID(IN:=#tCLEAN,L:=1,P:=#pos)) > 0 THEN
           (* charcter found skip to next one *)
           #pos := #pos + 1;
       ELSE
           (* wrong chracter needs to be deleted *)
           #tCLEAN := DELETE(IN:=#tCLEAN,L:=1,P:=#pos);
           #stop := #stop - 1;   (* the string is one character shorter now *)
       END_IF;
   END_WHILE;

   #CLEAN := #tCLEAN;


   (* revision history

   hm      18. jun. 2008   rev 1.0     
       original version 


   *)
END_FUNCTION

FUNCTION "CODE" : Byte   // FC229, SCL
TITLE = CODE
{ S7_Optimized_Access := 'FALSE' }
AUTHOR : hugo
FAMILY : STRINGS
NAME : CODE
VERSION : 1.1
// code extracts the code of a character at position POS of a string STR.
   VAR_INPUT
      STR : String[254];
      _STR AT STR : Struct
         length : Byte;
         act_length : Byte;
         str : Array[1..254] of Byte;
      END_STRUCT;
      POS : Int;
   END_VAR
   VAR_TEMP
      PT : Int;   // PT : POINTER TO BYTE;
   END_VAR
BEGIN


   IF #POS < 1 OR #POS > BYTE_TO_INT(#_STR.act_length) THEN
       #CODE := 0;
       RETURN;
   ELSE
       #PT := 1 + (#POS - 1);
       #CODE := #_STR.str[#PT];
   END_IF;

   (* revision history
   hm  9. mar. 2008    rev 1.0
       original version

   hm  29. mar. 2008   rev 1.1
       changed STRING to STRING(STRING_LENGTH)
   *)
END_FUNCTION

FUNCTION "COUNT_CHAR" : Int   // FC230, SCL
TITLE = COUNT_CHAR
{ S7_Optimized_Access := 'FALSE' }
AUTHOR : kurt
FAMILY : STRINGS
NAME : CT_CHR
VERSION : 1.1
// COUNT_CHAR how often a character CHAR occurs within a string STR.
   VAR_INPUT
      str : String[254];
      _str AT str : Struct
         length : Byte;
         act_length : Byte;
         str : Array[1..254] of Byte;
      END_STRUCT;
      chr : Byte;
   END_VAR
   VAR_TEMP
      l : Int;
      pt : Int;   // POINTER TO BYTE;
      pos : Int;
   END_VAR
BEGIN


   #pt := 1;                                //ADR(str);
   #l := BYTE_TO_INT(#_str.act_length);      //LEN(str);
   #COUNT_CHAR := 0;
   FOR #pos := 1 TO #l DO
       IF #_str.str[#pt] = #chr THEN #COUNT_CHAR := #COUNT_CHAR + 1; END_IF;
       #pt := #pt + 1;
   END_FOR;

   (* revision history
   hm  29. feb 2008    rev 1.0
       original version

   hm  29. mar. 2008   rev 1.1
       changed STRING to STRING(STRING_LENGTH)
   *)
END_FUNCTION

FUNCTION "DEC_TO_BYTE" : Byte   // FC231, SCL
TITLE = DEC_TO_BYTE
{ S7_Optimized_Access := 'FALSE' }
AUTHOR : hugo
FAMILY : STRINGS
NAME : DEC2BY
VERSION : 1.1
// DEC_TO_byte converts a decimal string into a byte.
   VAR_INPUT
      DEC : String[254];
      _DEC AT DEC : Struct
         length : Byte;
         act_length : Byte;
         str : Array[1..10] of Byte;
      END_STRUCT;
   END_VAR
   VAR_TEMP
      pt : Int;   // pt : POINTER TO BYTE;
      i : Int;
      X : Byte;
      stop : Int;
   END_VAR
BEGIN


   #pt := 1;        //ADR(dec);
   #stop := BYTE_TO_INT(#_DEC.act_length);    //LEN(DEC);
   FOR #i := 1 TO #stop DO
       (* read the first character and subtract 48 to get value in decimal 0 = 48 *)
       #X := #_DEC.str[#pt];
       (* calculate the value of the digit *)
       IF BYTE_TO_INT(#X) > 47 AND BYTE_TO_INT(#X) < 58 THEN
           #DEC_TO_BYTE := INT_TO_BYTE(BYTE_TO_INT(#DEC_TO_BYTE) * 10 + BYTE_TO_INT(#X) - 48);
       END_IF;
       #pt := #pt + 1;
   END_FOR;



   (* revision histroy
   hm  20. jun. 2008   rev 1.0
       original release

   hm  30. sep.2008    rev 1.1
       changed length of input string from 20 to 10
       corrected an error where decoding of characters 8 and 9 would fail

   *)
END_FUNCTION

FUNCTION "DEC_TO_DWORD" : DWord   // FC232, SCL
TITLE = DEC_TO_DWORD
{ S7_Optimized_Access := 'FALSE' }
AUTHOR : hugo
FAMILY : STRINGS
NAME : DEC2DW
VERSION : 1.1
// DEC_TO_DWORD converts a decimal string into a DWORD.
   VAR_INPUT
      DEC : String[254];
      _DEC AT DEC : Struct
         length : Byte;
         act_length : Byte;
         str : Array[1..20] of Byte;
      END_STRUCT;
   END_VAR
   VAR_TEMP
      pt : Int;   // pt : POINTER TO BYTE;
      i : Int;
      X : Byte;
      stop : Int;
   END_VAR
BEGIN


   #pt := 1;    //ADR(dec);
   #stop := BYTE_TO_INT(#_DEC.act_length);   //LEN(dec);
   FOR #i := 1 TO #stop DO
       (* read the first character and subtract 48 to get value in decimal 0 = 48 *)
       #X := #_DEC.str[#pt];
       (* calculate the value of the digit *)
       IF BYTE_TO_INT(#X) > 47 AND BYTE_TO_INT(#X) < 58 THEN
           #DEC_TO_DWORD := DINT_TO_DWORD(DWORD_TO_DINT(#DEC_TO_DWORD) * 10 + BYTE_TO_INT(#X) - 48);
       END_IF;
       #pt := #pt + 1;
   END_FOR;



   (* revision histroy
   hm  20. jun. 2008   rev 1.0
       original release

   hm  30. sep. 2008   rev 1.1
       corrected an error where decoding of characters 8 and 9 would fail
   *)
END_FUNCTION

FUNCTION "DEC_TO_INT" : Int   // FC233, SCL
TITLE = DEC_TO_INT
{ S7_Optimized_Access := 'FALSE' }
AUTHOR : hugo
FAMILY : STRINGS
NAME : DEC2INT
VERSION : 1.1
// DEC_TO_INT converts a decimal string into an Integer.
   VAR_INPUT
      DEC : String[254];
      _DEC AT DEC : Struct
         length : Byte;
         act_length : Byte;
         str : Array[1..10] of Byte;
      END_STRUCT;
   END_VAR
   VAR_TEMP
      pt : Int;   // pt : POINTER TO BYTE;
      i : Int;
      X : Byte;
      sign : Bool;
      stop : Int;
   END_VAR
BEGIN


   #pt := 1;    //ADR(dec);
   #stop := BYTE_TO_INT(#_DEC.act_length);   //LEN(dec);
   FOR #i := 1 TO #stop DO
       (* read the first character and subtract 48 to get value in decimal 0 = 48 *)
       #X := #_DEC.str[#pt];
       (* calculate the value of the digit *)
       IF BYTE_TO_INT(#X) > 47 AND BYTE_TO_INT(#X) < 58 THEN
           #DEC_TO_INT := #DEC_TO_INT * 10 + BYTE_TO_INT(#X) - 48;
       ELSIF #X = 45 AND #DEC_TO_INT = 0 THEN
           #sign := TRUE;
       END_IF;
       #pt := #pt + 1;
   END_FOR;
   IF #sign THEN #DEC_TO_INT := -#DEC_TO_INT; END_IF;


   (* revision histroy
   hm  20. jun. 2008   rev 1.0
       original release

   hm  30. sep. 2008   rev 1.1
       changed length of input string from 20 to 10
       corrected an error where decoding of characters 8 and 9 would fail
   *)
END_FUNCTION

FUNCTION "DEL_CHARS" : String[254]   // FC234, SCL
TITLE = DEL_CHARS
{ S7_Optimized_Access := 'FALSE' }
AUTHOR : hugo
FAMILY : STRINGS
NAME : DEL_CHR
VERSION : 1.0
// del_chars deletes all characters from a string which are specified in CX.
// 
// uses: LEN [FC21]
//       FIND [FC11]
//       MID [FC26]
//       DELETE [FC4]
   VAR_INPUT
      IN : String[254];
      CX : String[254];
   END_VAR
   VAR_TEMP
      tDEL_CHARS : String[254];
      tCX : String[80];
      pos : Int;
      stop : Int;
   END_VAR
BEGIN


   #pos := 1;
   #tDEL_CHARS := #IN;
   #tCX := #CX;

   (* copy input string *)
   //DEL_CHARS := IN;
   #stop := LEN(#tDEL_CHARS);
   WHILE #pos <= #stop DO
       IF FIND(IN1:=#tCX,IN2:=MID(IN:=#tDEL_CHARS,L:=1,P:=#pos)) > 0 THEN
           (* wrong chracter needs to be deleted *)
           #tDEL_CHARS := DELETE(IN:=#tDEL_CHARS,L:=1,P:=#pos);
           #stop := #stop - 1;   (* the string is one character shorter now *)
       ELSE
           (* charcter not found skip to next one *)
           #pos := #pos + 1;
       END_IF;
   END_WHILE;

   #DEL_CHARS := #tDEL_CHARS;


   (* revision history

   hm      18. jun. 2008   rev 1.0     
       original version 


   *)
END_FUNCTION

FUNCTION "DT_TO_STRF" : String[254]   // FC235, SCL
TITLE = DT_TO_STRF
{ S7_Optimized_Access := 'FALSE' }
AUTHOR : hugo
FAMILY : STRINGS
NAME : DT2STRF
VERSION : 1.1
// DT_TO_STRINGF converts a DATETIME input to a formatted string
// 
// uses: LANGUAGE [DB4]
//       I_STRNG [FC16]
//       CONCAT [FC2]
//       DT_DATE [FC6]
//       DT_TOD [FC8]
//       FIND [FC11]
//       CODE [FC229]
//       DELETE [FC4]
//       YEAR_OF_DATE [FC219]
//       RIGHT [FC32]
//       MONTH_OF_DATE [FC202]
//       DAY_OF_YEAR [FC180] 
//       YEAR_BEGIN [FC217]
//       LEAP_OF_DATE [FC193] 
//       LEAP_YEAR [FC194]
//       LEN [FC21]
//       MONTH_TO_STRING [FC275]
//       DAY_OF_MONTH [FC178]
//       DAY_OF_WEEK [FC179]
//       WEEKDAY_TO_STRING [FC289]
//       HOUR [FC187]
//       MINUTE [FC197]
//       SECOND [FC210]
//       REPLACE [FC31]
   VAR_INPUT
      DTI : Date_And_Time;
      MS : Int;
      FMT : String[254];
      LANG : Int;
   END_VAR
   VAR_TEMP
      tDT_TO_STRF : String[254];
      _DT_TO_STRF AT tDT_TO_STRF : Struct
         length : Byte;
         act_length : Byte;
         str : Array[1..254] of Byte;
      END_STRUCT;
      tDTI : Date_And_Time;
      ly : Int;
      dx : Date;
      fs : String[10];
      td : Time_Of_Day;
      tmp : Int;
      pos : Int;
      f : Int;
   END_VAR
BEGIN


   IF #LANG < 1 THEN #ly := "LANGUAGE".DEFAULT; ELSE #ly := MIN(IN1:="LANGUAGE".LMAX, IN2:=#LANG); END_IF;

   (* decode date and time information *)
   #tDTI := #DTI;
   #dx := T_CONV(#tDTI);
   #td := T_CONV(#tDTI);